REGION Network 20: Total Time Machine
   // ENO of a box is taken as its EN; it also drops when the box reports an error
   "Data_TimeData"."Total Time Machine" := "Data_TimeData"."Mesin Run" + "Data_TimeData"."Mesin Run Baypass" + "Data_TimeData"."Mesin Stop" + "Data_TimeData"."Mesin Error";
   "Data_TODData"."Total Time Machine" := T_CONV(IN := "Data_TimeData"."Total Time Machine");
   "Data_DTLData"."Total Time Machine"[0] := T_COMBINE(IN1 := D#1990-01-01,
                           IN2 := "Data_TODData"."Total Time Machine");
END_REGION

REGION Network 21: % Persen Counter Mesin Terhadap Lama Current Shift
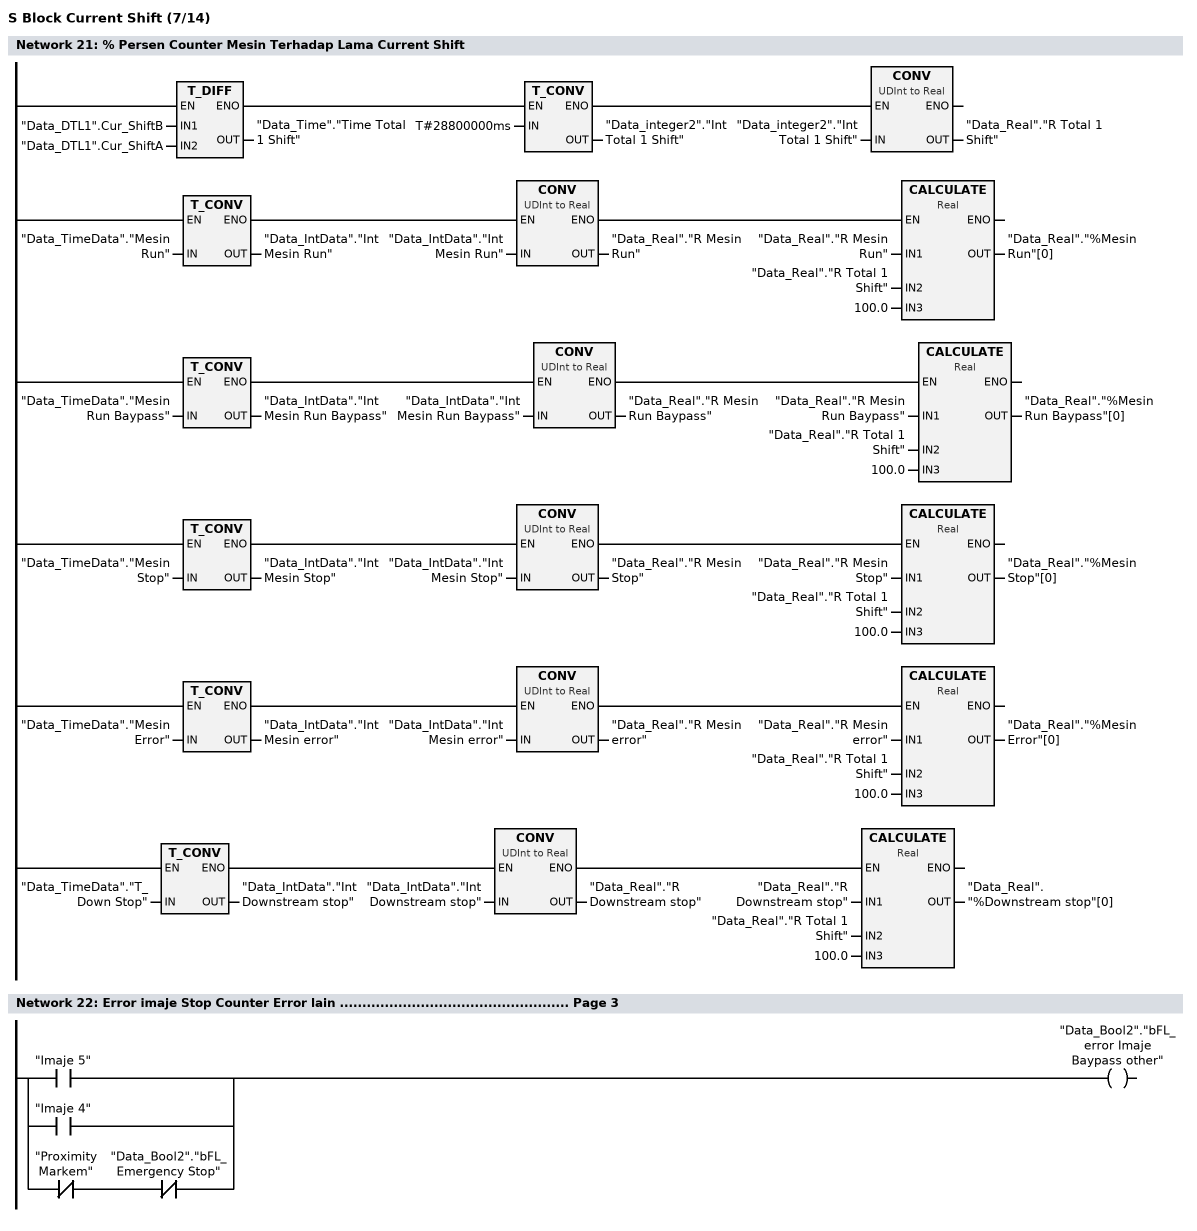
   // ENO of a box is taken as its EN; it also drops when the box reports an error
   "Data_Time"."Time Total 1 Shift" := T_DIFF(IN1 := "Data_DTL1".Cur_ShiftB, IN2 := "Data_DTL1".Cur_ShiftA);
   "Data_integer2"."Int Total 1 Shift" := T_CONV(IN := T#28800000ms);
   "Data_Real"."R Total 1 Shift" := UDINT_TO_REAL("Data_integer2"."Int Total 1 Shift");
   "Data_IntData"."Int Mesin Run" := T_CONV(IN := "Data_TimeData"."Mesin Run");
   "Data_Real"."R Mesin Run" := UDINT_TO_REAL("Data_IntData"."Int Mesin Run");
   "Data_Real"."%Mesin Run"[0] := ("Data_Real"."R Mesin Run"/"Data_Real"."R Total 1 Shift")*100.0;
   "Data_IntData"."Int Mesin Run Baypass" := T_CONV(IN := "Data_TimeData"."Mesin Run Baypass");
   "Data_Real"."R Mesin Run Baypass" := UDINT_TO_REAL("Data_IntData"."Int Mesin Run Baypass");
   "Data_Real"."%Mesin Run Baypass"[0] := ("Data_Real"."R Mesin Run Baypass"/"Data_Real"."R Total 1 Shift")*100.0;
   "Data_IntData"."Int Mesin Stop" := T_CONV(IN := "Data_TimeData"."Mesin Stop");
   "Data_Real"."R Mesin Stop" := UDINT_TO_REAL("Data_IntData"."Int Mesin Stop");
   "Data_Real"."%Mesin Stop"[0] := ("Data_Real"."R Mesin Stop"/"Data_Real"."R Total 1 Shift")*100.0;
   "Data_IntData"."Int Mesin error" := T_CONV(IN := "Data_TimeData"."Mesin Error");
   "Data_Real"."R Mesin error" := UDINT_TO_REAL("Data_IntData"."Int Mesin error");
   "Data_Real"."%Mesin Error"[0] := ("Data_Real"."R Mesin error"/"Data_Real"."R Total 1 Shift")*100.0;
   "Data_IntData"."Int Downstream stop" := T_CONV(IN := "Data_TimeData"."T_Down Stop");
   "Data_Real"."R Downstream stop" := UDINT_TO_REAL("Data_IntData"."Int Downstream stop");
   "Data_Real"."%Downstream stop"[0] := ("Data_Real"."R Downstream stop"/"Data_Real"."R Total 1 Shift")*100.0;
END_REGION

REGION Network 22: Error imaje Stop Counter Error lain ................................................... Page 3
   RUNG wire#powerrail
      Contact( "Imaje 5" )
      wire#w1
      Coil( "Data_Bool2"."bFL_error Imaje Baypass other" )
   END_RUNG
   RUNG wire#powerrail
      Contact( "Imaje 4" )
   END_RUNG wire#w1
   RUNG wire#powerrail
      I_Contact( "Proximity Markem" )
      I_Contact( "Data_Bool2"."bFL_Emergency Stop" )
   END_RUNG wire#w1
   // the same network as SCL:
   "Data_Bool2"."bFL_error Imaje Baypass other" := "Imaje 5" OR "Imaje 4" OR (NOT "Proximity Markem" AND NOT "Data_Bool2"."bFL_Emergency Stop");
END_REGION

REGION Network 23: 1. Counter Imaje System Error
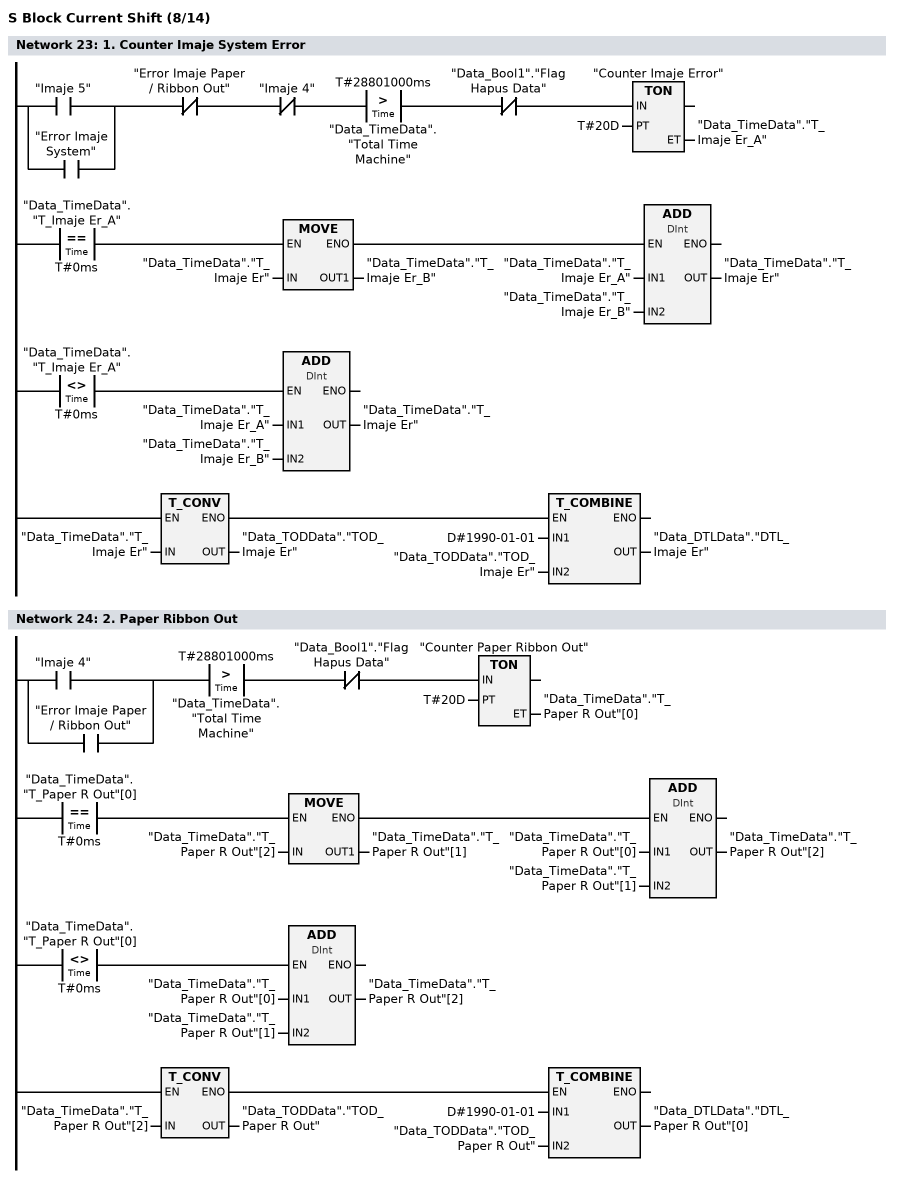
   // ENO of a box is taken as its EN; it also drops when the box reports an error
   "Counter Imaje Error".TON(IN := ("Imaje 5" OR "Error Imaje System") AND NOT "Error Imaje Paper / Ribbon Out" AND NOT "Imaje 4" AND (T#28801000ms > "Data_TimeData"."Total Time Machine") AND NOT "Data_Bool1"."Flag Hapus Data",
                           PT := T#20D,
                           ET => "Data_TimeData"."T_Imaje Er_A");
   IF "Data_TimeData"."T_Imaje Er_A" = T#0ms THEN
       "Data_TimeData"."T_Imaje Er_B" := "Data_TimeData"."T_Imaje Er";
       "Data_TimeData"."T_Imaje Er" := "Data_TimeData"."T_Imaje Er_A" + "Data_TimeData"."T_Imaje Er_B";
   END_IF;
   IF "Data_TimeData"."T_Imaje Er_A" <> T#0ms THEN
       "Data_TimeData"."T_Imaje Er" := "Data_TimeData"."T_Imaje Er_A" + "Data_TimeData"."T_Imaje Er_B";
   END_IF;
   "Data_TODData"."TOD_Imaje Er" := T_CONV(IN := "Data_TimeData"."T_Imaje Er");
   "Data_DTLData"."DTL_Imaje Er" := T_COMBINE(IN1 := D#1990-01-01, IN2 := "Data_TODData"."TOD_Imaje Er");
END_REGION

REGION Network 24: 2. Paper Ribbon Out
   // ENO of a box is taken as its EN; it also drops when the box reports an error
   "Counter Paper Ribbon Out".TON(IN := ("Imaje 4" OR "Error Imaje Paper / Ribbon Out") AND (T#28801000ms > "Data_TimeData"."Total Time Machine") AND NOT "Data_Bool1"."Flag Hapus Data",
                           PT := T#20D,
                           ET => "Data_TimeData"."T_Paper R Out"[0]);
   #_w1 := "Data_TimeData"."T_Paper R Out"[0] = T#0ms;
   IF #_w1 THEN
       "Data_TimeData"."T_Paper R Out"[1] := "Data_TimeData"."T_Paper R Out"[2];
       "Data_TimeData"."T_Paper R Out"[2] := "Data_TimeData"."T_Paper R Out"[0] + "Data_TimeData"."T_Paper R Out"[1];
   END_IF;
   IF "Data_TimeData"."T_Paper R Out"[0] <> T#0ms THEN
       "Data_TimeData"."T_Paper R Out"[2] := "Data_TimeData"."T_Paper R Out"[0] + "Data_TimeData"."T_Paper R Out"[1];
   END_IF;
   "Data_TODData"."TOD_Paper R Out" := T_CONV(IN := "Data_TimeData"."T_Paper R Out"[2]);
   "Data_DTLData"."DTL_Paper R Out"[0] := T_COMBINE(IN1 := D#1990-01-01,
                           IN2 := "Data_TODData"."TOD_Paper R Out");
END_REGION

REGION Network 25: 3. Imaje Not In Position
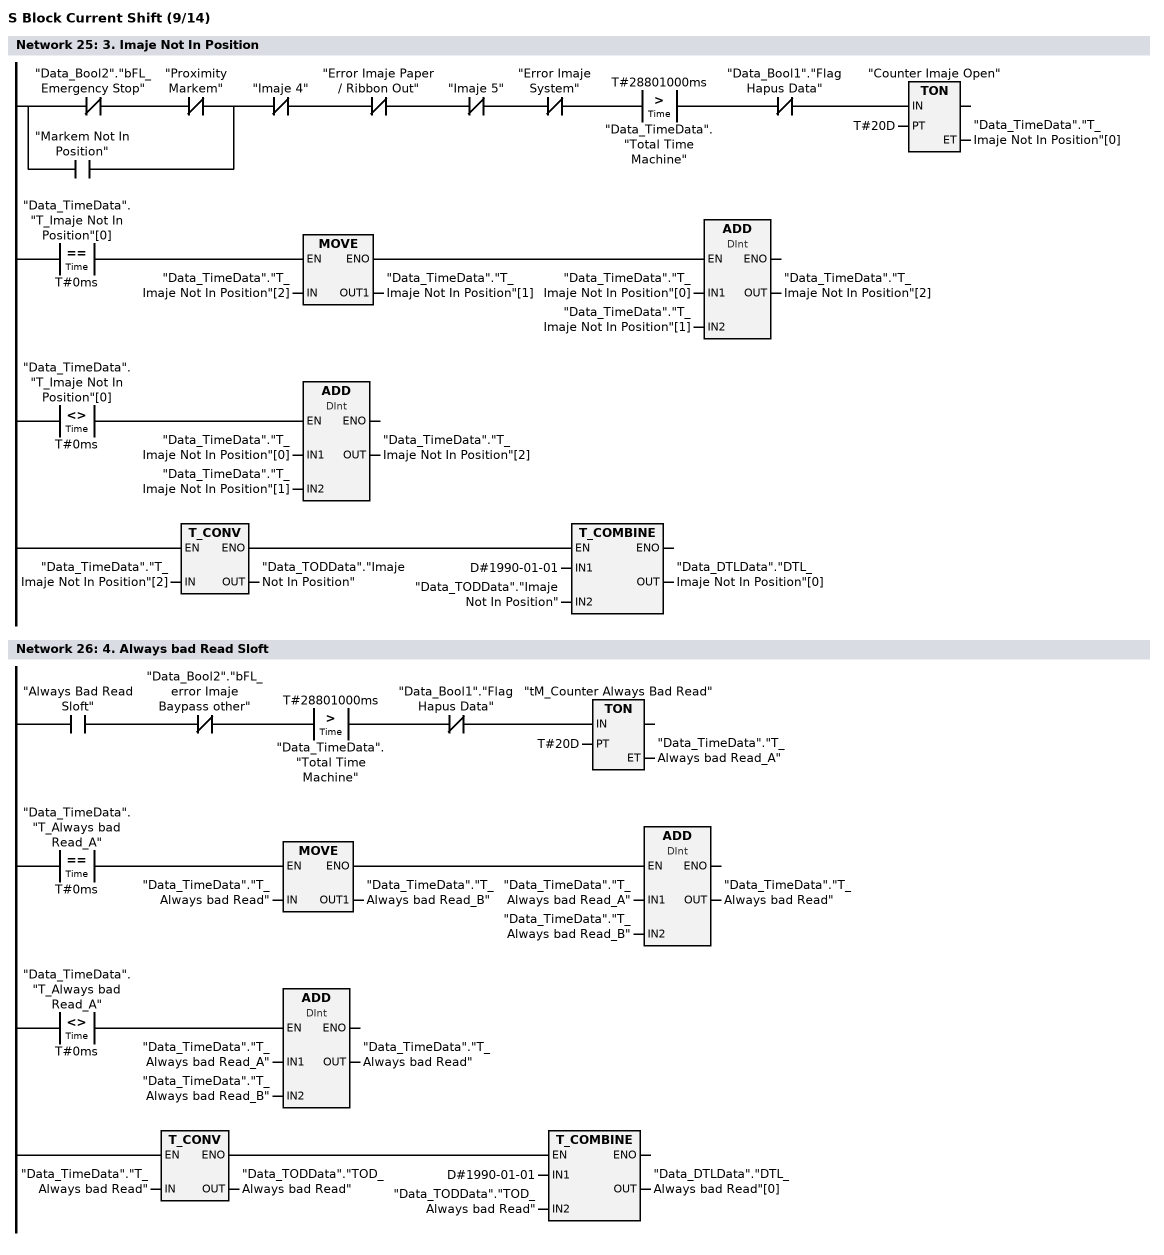
   // ENO of a box is taken as its EN; it also drops when the box reports an error
   "Counter Imaje Open".TON(IN := ((NOT "Data_Bool2"."bFL_Emergency Stop" AND NOT "Proximity Markem") OR "Markem Not In Position") AND NOT "Imaje 4" AND NOT "Error Imaje Paper / Ribbon Out" AND NOT "Imaje 5" AND NOT "Error Imaje System" AND (T#28801000ms > "Data_TimeData"."Total Time Machine") AND NOT "Data_Bool1"."Flag Hapus Data",
                           PT := T#20D,
                           ET => "Data_TimeData"."T_Imaje Not In Position"[0]);
   #_w1 := "Data_TimeData"."T_Imaje Not In Position"[0] = T#0ms;
   IF #_w1 THEN
       "Data_TimeData"."T_Imaje Not In Position"[1] := "Data_TimeData"."T_Imaje Not In Position"[2];
       "Data_TimeData"."T_Imaje Not In Position"[2] := "Data_TimeData"."T_Imaje Not In Position"[0] + "Data_TimeData"."T_Imaje Not In Position"[1];
   END_IF;
   IF "Data_TimeData"."T_Imaje Not In Position"[0] <> T#0ms THEN
       "Data_TimeData"."T_Imaje Not In Position"[2] := "Data_TimeData"."T_Imaje Not In Position"[0] + "Data_TimeData"."T_Imaje Not In Position"[1];
   END_IF;
   "Data_TODData"."Imaje Not In Position" := T_CONV(IN := "Data_TimeData"."T_Imaje Not In Position"[2]);
   "Data_DTLData"."DTL_Imaje Not In Position"[0] := T_COMBINE(IN1 := D#1990-01-01,
                           IN2 := "Data_TODData"."Imaje Not In Position");
END_REGION

REGION Network 26: 4. Always bad Read Sloft
   // ENO of a box is taken as its EN; it also drops when the box reports an error
   "tM_Counter Always Bad Read".TON(IN := "Always Bad Read Sloft" AND NOT "Data_Bool2"."bFL_error Imaje Baypass other" AND (T#28801000ms > "Data_TimeData"."Total Time Machine") AND NOT "Data_Bool1"."Flag Hapus Data",
                           PT := T#20D,
                           ET => "Data_TimeData"."T_Always bad Read_A");
   IF "Data_TimeData"."T_Always bad Read_A" = T#0ms THEN
       "Data_TimeData"."T_Always bad Read_B" := "Data_TimeData"."T_Always bad Read";
       "Data_TimeData"."T_Always bad Read" := "Data_TimeData"."T_Always bad Read_A" + "Data_TimeData"."T_Always bad Read_B";
   END_IF;
   IF "Data_TimeData"."T_Always bad Read_A" <> T#0ms THEN
       "Data_TimeData"."T_Always bad Read" := "Data_TimeData"."T_Always bad Read_A" + "Data_TimeData"."T_Always bad Read_B";
   END_IF;
   "Data_TODData"."TOD_Always bad Read" := T_CONV(IN := "Data_TimeData"."T_Always bad Read");
   "Data_DTLData"."DTL_Always bad Read"[0] := T_COMBINE(IN1 := D#1990-01-01,
                           IN2 := "Data_TODData"."TOD_Always bad Read");
END_REGION

REGION Network 27: 5. Counter Sloft Jammed
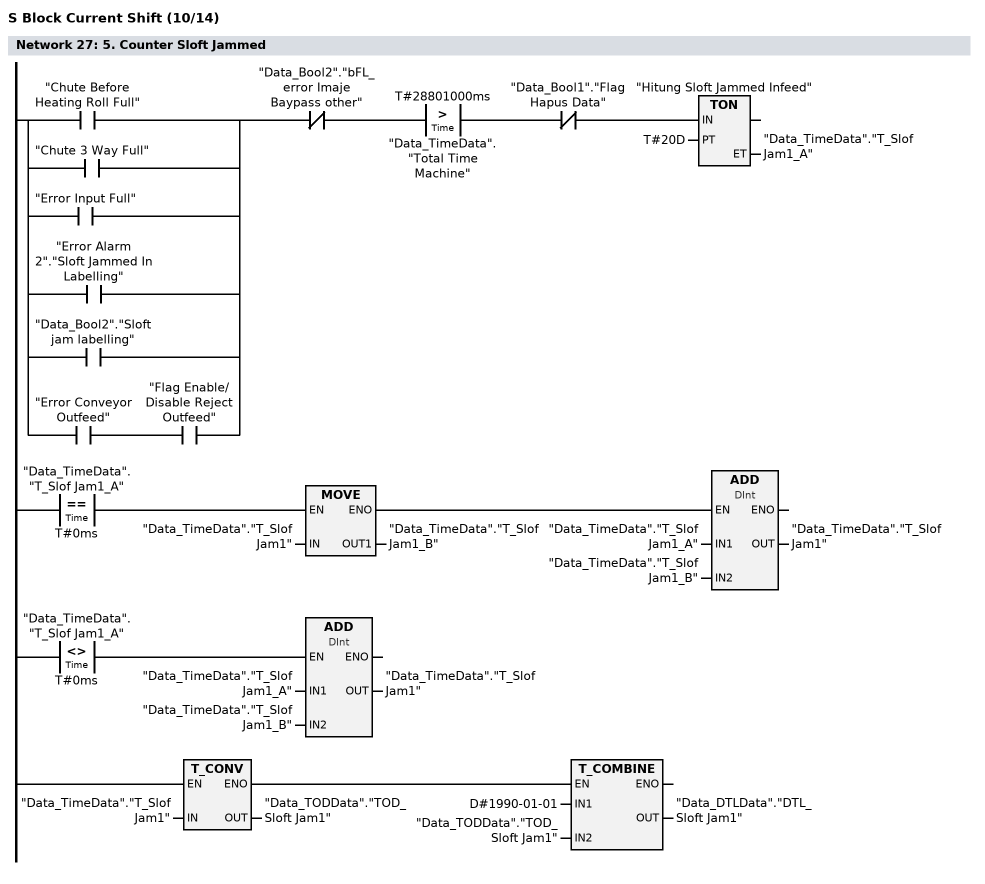
   // ENO of a box is taken as its EN; it also drops when the box reports an error
   "Hitung Sloft Jammed Infeed".TON(IN := ("Chute Before Heating Roll Full" OR "Chute 3 Way Full" OR "Error Input Full" OR "Error Alarm 2"."Sloft Jammed In Labelling" OR "Data_Bool2"."Sloft jam labelling" OR ("Error Conveyor Outfeed" AND "Flag Enable/Disable Reject Outfeed")) AND NOT "Data_Bool2"."bFL_error Imaje Baypass other" AND (T#28801000ms > "Data_TimeData"."Total Time Machine") AND NOT "Data_Bool1"."Flag Hapus Data",
                           PT := T#20D,
                           ET => "Data_TimeData"."T_Slof Jam1_A");
   IF "Data_TimeData"."T_Slof Jam1_A" = T#0ms THEN
       "Data_TimeData"."T_Slof Jam1_B" := "Data_TimeData"."T_Slof Jam1";
       "Data_TimeData"."T_Slof Jam1" := "Data_TimeData"."T_Slof Jam1_A" + "Data_TimeData"."T_Slof Jam1_B";
   END_IF;
   IF "Data_TimeData"."T_Slof Jam1_A" <> T#0ms THEN
       "Data_TimeData"."T_Slof Jam1" := "Data_TimeData"."T_Slof Jam1_A" + "Data_TimeData"."T_Slof Jam1_B";
   END_IF;
   "Data_TODData"."TOD_Sloft Jam1" := T_CONV(IN := "Data_TimeData"."T_Slof Jam1");
   "Data_DTLData"."DTL_Sloft Jam1" := T_COMBINE(IN1 := D#1990-01-01, IN2 := "Data_TODData"."TOD_Sloft Jam1");
END_REGION

REGION Network 28: 6. Counter Pressure Low
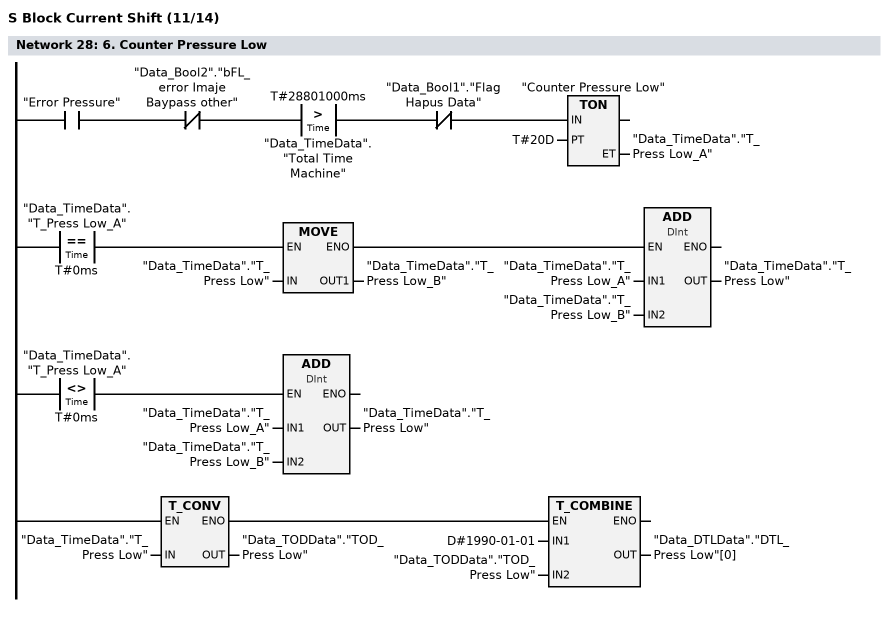
   // ENO of a box is taken as its EN; it also drops when the box reports an error
   "Counter Pressure Low".TON(IN := "Error Pressure" AND NOT "Data_Bool2"."bFL_error Imaje Baypass other" AND (T#28801000ms > "Data_TimeData"."Total Time Machine") AND NOT "Data_Bool1"."Flag Hapus Data",
                           PT := T#20D,
                           ET => "Data_TimeData"."T_Press Low_A");
   IF "Data_TimeData"."T_Press Low_A" = T#0ms THEN
       "Data_TimeData"."T_Press Low_B" := "Data_TimeData"."T_Press Low";
       "Data_TimeData"."T_Press Low" := "Data_TimeData"."T_Press Low_A" + "Data_TimeData"."T_Press Low_B";
   END_IF;
   IF "Data_TimeData"."T_Press Low_A" <> T#0ms THEN
       "Data_TimeData"."T_Press Low" := "Data_TimeData"."T_Press Low_A" + "Data_TimeData"."T_Press Low_B";
   END_IF;
   "Data_TODData"."TOD_Press Low" := T_CONV(IN := "Data_TimeData"."T_Press Low");
   "Data_DTLData"."DTL_Press Low"[0] := T_COMBINE(IN1 := D#1990-01-01, IN2 := "Data_TODData"."TOD_Press Low");
END_REGION

REGION Network 29: 7. Counter RS Pneumatic Error
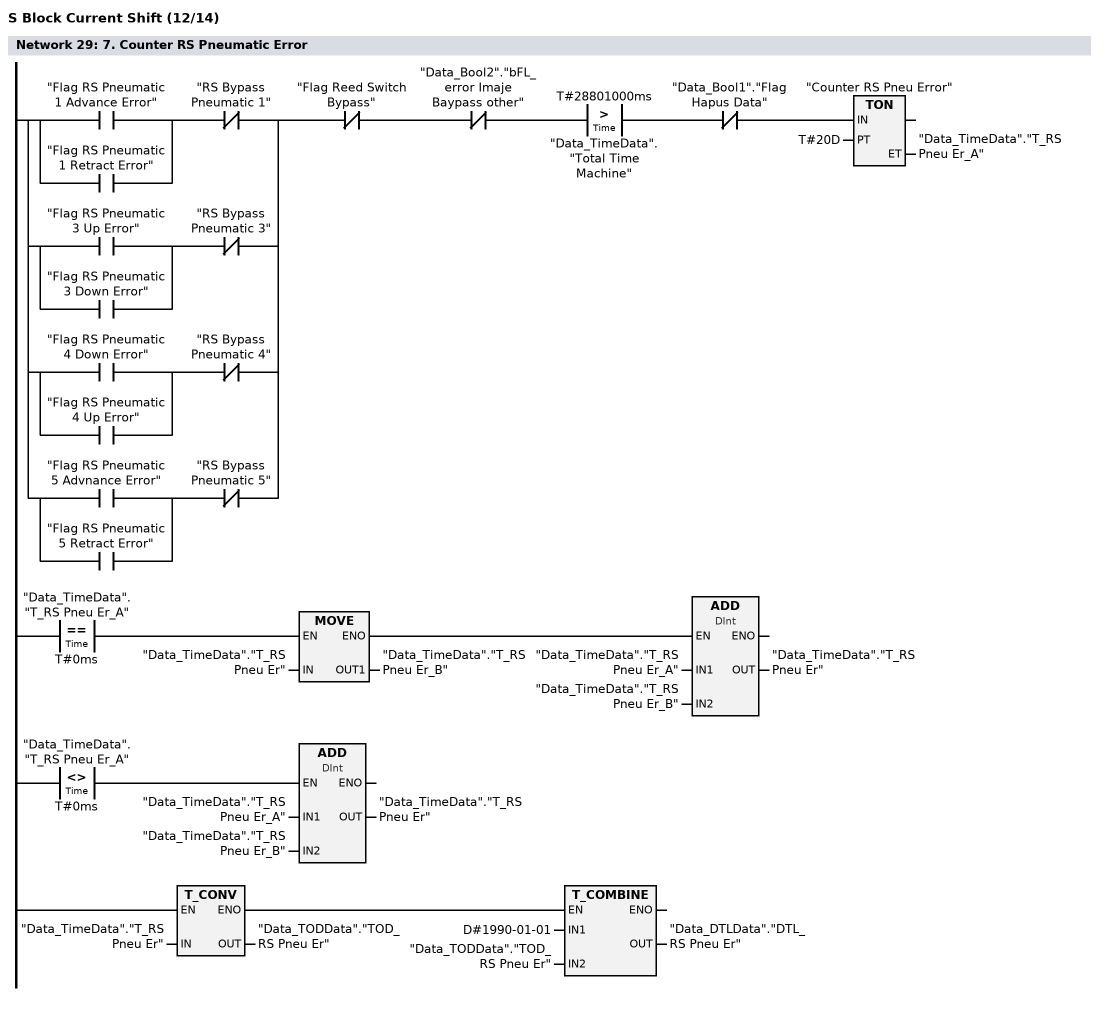
   // ENO of a box is taken as its EN; it also drops when the box reports an error
   "Counter RS Pneu Error".TON(IN := ((("Flag RS Pneumatic 1 Advance Error" OR "Flag RS Pneumatic 1 Retract Error") AND NOT "RS Bypass Pneumatic 1") OR (("Flag RS Pneumatic 3 Up Error" OR "Flag RS Pneumatic 3 Down Error") AND NOT "RS Bypass Pneumatic 3") OR (("Flag RS Pneumatic 4 Down Error" OR "Flag RS Pneumatic 4 Up Error") AND NOT "RS Bypass Pneumatic 4") OR (("Flag RS Pneumatic 5 Advnance Error" OR "Flag RS Pneumatic 5 Retract Error") AND NOT "RS Bypass Pneumatic 5")) AND NOT "Flag Reed Switch Bypass" AND NOT "Data_Bool2"."bFL_error Imaje Baypass other" AND (T#28801000ms > "Data_TimeData"."Total Time Machine") AND NOT "Data_Bool1"."Flag Hapus Data",
                           PT := T#20D,
                           ET => "Data_TimeData"."T_RS Pneu Er_A");
   IF "Data_TimeData"."T_RS Pneu Er_A" = T#0ms THEN
       "Data_TimeData"."T_RS Pneu Er_B" := "Data_TimeData"."T_RS Pneu Er";
       "Data_TimeData"."T_RS Pneu Er" := "Data_TimeData"."T_RS Pneu Er_A" + "Data_TimeData"."T_RS Pneu Er_B";
   END_IF;
   IF "Data_TimeData"."T_RS Pneu Er_A" <> T#0ms THEN
       "Data_TimeData"."T_RS Pneu Er" := "Data_TimeData"."T_RS Pneu Er_A" + "Data_TimeData"."T_RS Pneu Er_B";
   END_IF;
   "Data_TODData"."TOD_RS Pneu Er" := T_CONV(IN := "Data_TimeData"."T_RS Pneu Er");
   "Data_DTLData"."DTL_RS Pneu Er" := T_COMBINE(IN1 := D#1990-01-01, IN2 := "Data_TODData"."TOD_RS Pneu Er");
END_REGION

REGION Network 30: 8. Counter Door open error
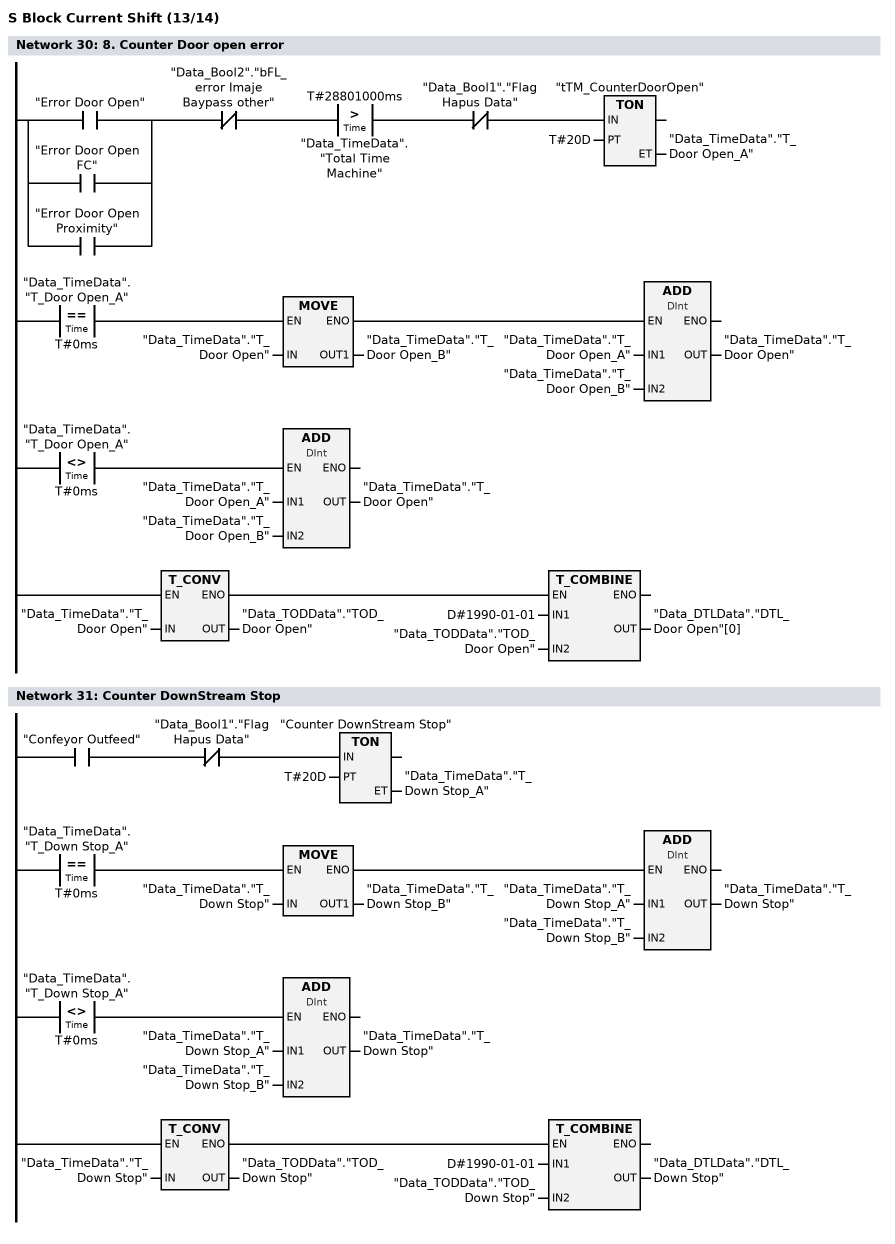
   // ENO of a box is taken as its EN; it also drops when the box reports an error
   "tTM_CounterDoorOpen".TON(IN := ("Error Door Open" OR "Error Door Open FC" OR "Error Door Open Proximity") AND NOT "Data_Bool2"."bFL_error Imaje Baypass other" AND (T#28801000ms > "Data_TimeData"."Total Time Machine") AND NOT "Data_Bool1"."Flag Hapus Data",
                           PT := T#20D,
                           ET => "Data_TimeData"."T_Door Open_A");
   IF "Data_TimeData"."T_Door Open_A" = T#0ms THEN
       "Data_TimeData"."T_Door Open_B" := "Data_TimeData"."T_Door Open";
       "Data_TimeData"."T_Door Open" := "Data_TimeData"."T_Door Open_A" + "Data_TimeData"."T_Door Open_B";
   END_IF;
   IF "Data_TimeData"."T_Door Open_A" <> T#0ms THEN
       "Data_TimeData"."T_Door Open" := "Data_TimeData"."T_Door Open_A" + "Data_TimeData"."T_Door Open_B";
   END_IF;
   "Data_TODData"."TOD_Door Open" := T_CONV(IN := "Data_TimeData"."T_Door Open");
   "Data_DTLData"."DTL_Door Open"[0] := T_COMBINE(IN1 := D#1990-01-01, IN2 := "Data_TODData"."TOD_Door Open");
END_REGION

REGION Network 31: Counter DownStream Stop
   // ENO of a box is taken as its EN; it also drops when the box reports an error
   "Counter DownStream Stop".TON(IN := "Confeyor Outfeed" AND NOT "Data_Bool1"."Flag Hapus Data",
                           PT := T#20D,
                           ET => "Data_TimeData"."T_Down Stop_A");
   IF "Data_TimeData"."T_Down Stop_A" = T#0ms THEN
       "Data_TimeData"."T_Down Stop_B" := "Data_TimeData"."T_Down Stop";
       "Data_TimeData"."T_Down Stop" := "Data_TimeData"."T_Down Stop_A" + "Data_TimeData"."T_Down Stop_B";
   END_IF;
   IF "Data_TimeData"."T_Down Stop_A" <> T#0ms THEN
       "Data_TimeData"."T_Down Stop" := "Data_TimeData"."T_Down Stop_A" + "Data_TimeData"."T_Down Stop_B";
   END_IF;
   "Data_TODData"."TOD_Down Stop" := T_CONV(IN := "Data_TimeData"."T_Down Stop");
   "Data_DTLData"."DTL_Down Stop" := T_COMBINE(IN1 := D#1990-01-01, IN2 := "Data_TODData"."TOD_Down Stop");
END_REGION

REGION Network 32: Total Error
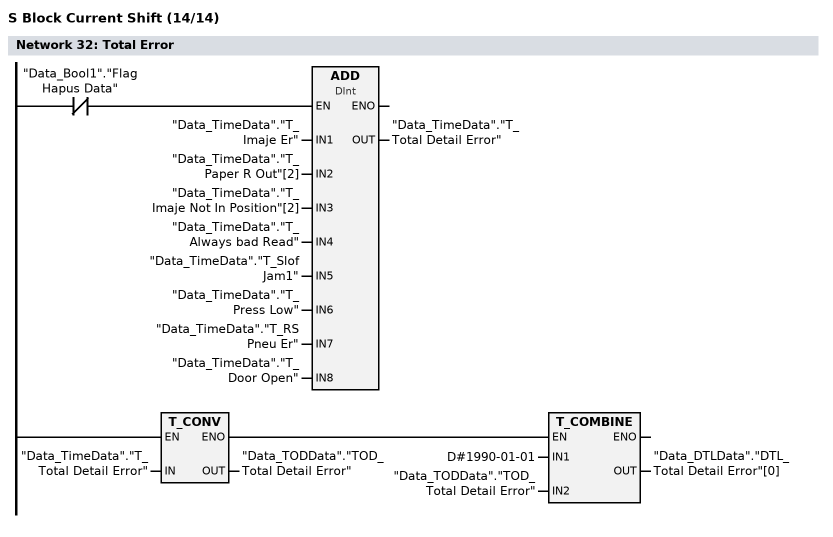
   // ENO of a box is taken as its EN; it also drops when the box reports an error
   IF NOT "Data_Bool1"."Flag Hapus Data" THEN
       "Data_TimeData"."T_Total Detail Error" := "Data_TimeData"."T_Imaje Er" + "Data_TimeData"."T_Paper R Out"[2] + "Data_TimeData"."T_Imaje Not In Position"[2] + "Data_TimeData"."T_Always bad Read" + "Data_TimeData"."T_Slof Jam1" + "Data_TimeData"."T_Press Low" + "Data_TimeData"."T_RS Pneu Er" + "Data_TimeData"."T_Door Open";
   END_IF;
   "Data_TODData"."TOD_Total Detail Error" := T_CONV(IN := "Data_TimeData"."T_Total Detail Error");
   "Data_DTLData"."DTL_Total Detail Error"[0] := T_COMBINE(IN1 := D#1990-01-01,
                           IN2 := "Data_TODData"."TOD_Total Detail Error");
END_REGION
END_FUNCTION_BLOCK

FUNCTION_BLOCK "Block Labeling"   // FB5, LAD
{ S7_Optimized_Access := 'TRUE' }
VERSION : 0.1
   VAR_TEMP   // added for the SCL form of the ladder/FBD networks
      _w1 : Bool;
      _w2 : Bool;
      _w3 : Bool;
      _w4 : Bool;
   END_VAR
BEGIN

REGION Network 1: By pass ON
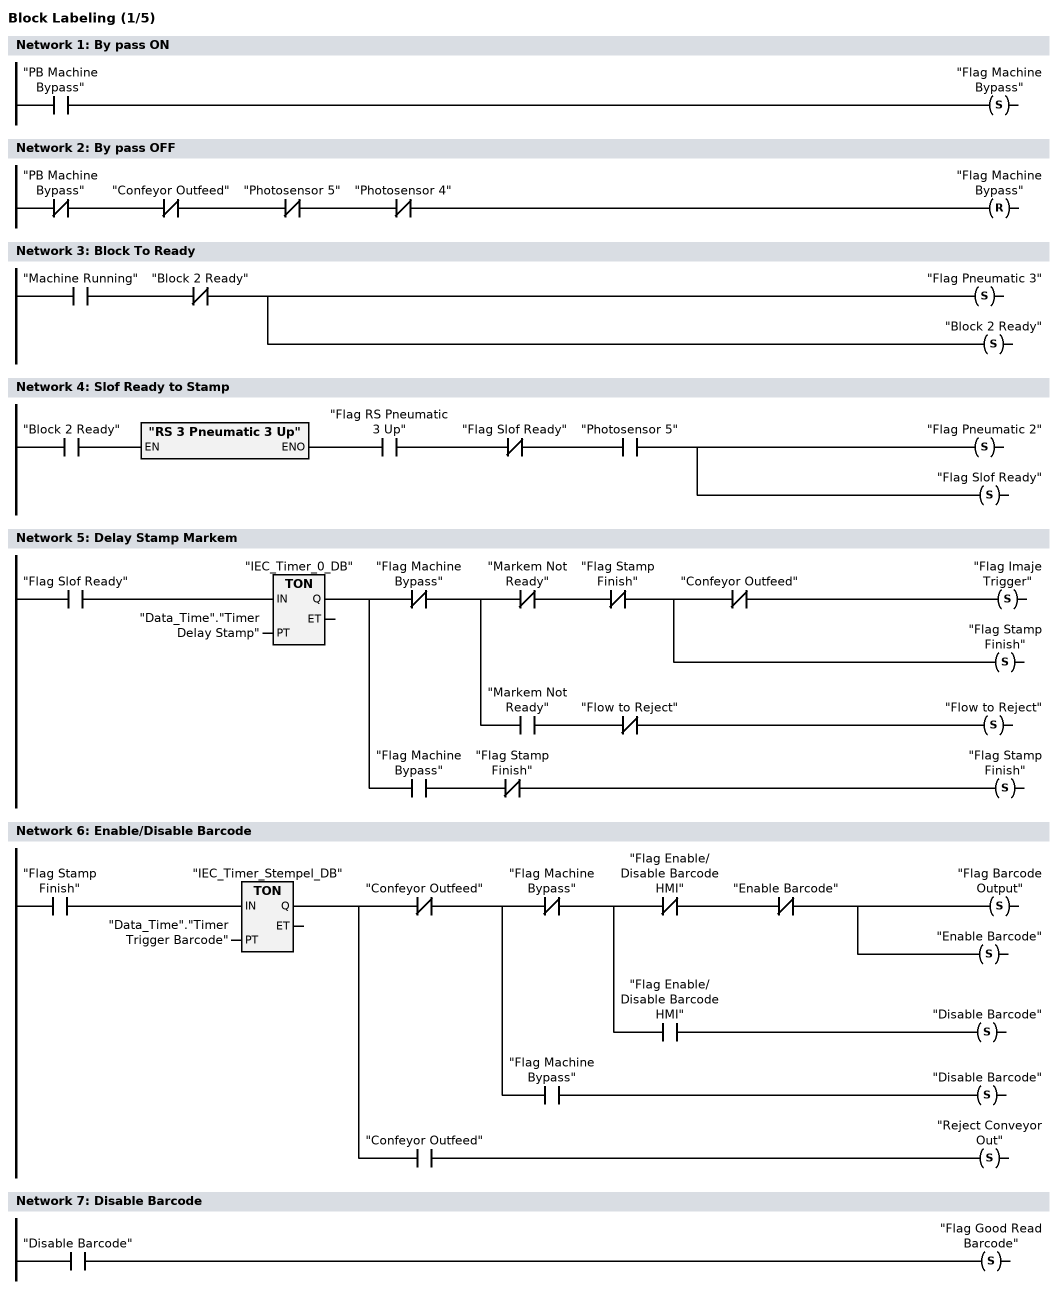
   RUNG wire#powerrail
      Contact( "PB Machine Bypass" )
      S_Coil( "Flag Machine Bypass" )
   END_RUNG
   // the same network as SCL:
   IF "PB Machine Bypass" THEN "Flag Machine Bypass" := TRUE; END_IF;
END_REGION

REGION Network 2: By pass OFF
   RUNG wire#powerrail
      I_Contact( "PB Machine Bypass" )
      I_Contact( "Confeyor Outfeed" )
      I_Contact( "Photosensor 5" )
      I_Contact( "Photosensor 4" )
      R_Coil( "Flag Machine Bypass" )
   END_RUNG
   // the same network as SCL:
   IF NOT "PB Machine Bypass" AND NOT "Confeyor Outfeed" AND NOT "Photosensor 5" AND NOT "Photosensor 4" THEN
       "Flag Machine Bypass" := FALSE;
   END_IF;
END_REGION

REGION Network 3: Block To Ready
   RUNG wire#powerrail
      Contact( "Machine Running" )
      I_Contact( "Block 2 Ready" )
      wire#w1
      S_Coil( "Flag Pneumatic 3" )
   END_RUNG
   RUNG wire#w1
      S_Coil( "Block 2 Ready" )
   END_RUNG
   // the same network as SCL:
   IF "Machine Running" AND NOT "Block 2 Ready" THEN
       "Flag Pneumatic 3" := TRUE;
       "Block 2 Ready" := TRUE;
   END_IF;
END_REGION

REGION Network 4: Slof Ready to Stamp
   RUNG wire#powerrail
      Contact( "Block 2 Ready" )
      "RS 3 Pneumatic 3 Up"()
      Contact( "Flag RS Pneumatic 3 Up" )
      I_Contact( "Flag Slof Ready" )
      Contact( "Photosensor 5" )
      wire#w1
      S_Coil( "Flag Pneumatic 2" )
   END_RUNG
   RUNG wire#w1
      S_Coil( "Flag Slof Ready" )
   END_RUNG
   // the same network as SCL:
   "RS 3 Pneumatic 3 Up"(EN := "Block 2 Ready", ENO => #_w1);
   IF #_w1 AND "Flag RS Pneumatic 3 Up" AND NOT "Flag Slof Ready" AND "Photosensor 5" THEN
       "Flag Pneumatic 2" := TRUE;
       "Flag Slof Ready" := TRUE;
   END_IF;
END_REGION

REGION Network 5: Delay Stamp Markem
   "IEC_Timer_0_DB".TON(IN := "Flag Slof Ready", PT := "Data_Time"."Timer Delay Stamp");
   #_w1 := "IEC_Timer_0_DB".Q AND NOT "Flag Machine Bypass";
   #_w2 := #_w1 AND NOT "Markem Not Ready" AND NOT "Flag Stamp Finish";
   IF #_w2 AND NOT "Confeyor Outfeed" THEN "Flag Imaje Trigger" := TRUE; END_IF;
   IF #_w2 THEN "Flag Stamp Finish" := TRUE; END_IF;
   IF #_w1 AND "Markem Not Ready" AND NOT "Flow to Reject" THEN "Flow to Reject" := TRUE; END_IF;
   IF "IEC_Timer_0_DB".Q AND "Flag Machine Bypass" AND NOT "Flag Stamp Finish" THEN
       "Flag Stamp Finish" := TRUE;
   END_IF;
END_REGION

REGION Network 6: Enable/Disable Barcode
   "IEC_Timer_Stempel_DB".TON(IN := "Flag Stamp Finish", PT := "Data_Time"."Timer Trigger Barcode");
   #_w1 := "IEC_Timer_Stempel_DB".Q AND NOT "Confeyor Outfeed";
   #_w2 := #_w1 AND NOT "Flag Machine Bypass";
   IF #_w2 AND NOT "Flag Enable/Disable Barcode HMI" AND NOT "Enable Barcode" THEN
       "Flag Barcode Output" := TRUE;
       "Enable Barcode" := TRUE;
   END_IF;
   IF #_w2 AND "Flag Enable/Disable Barcode HMI" THEN "Disable Barcode" := TRUE; END_IF;
   IF #_w1 AND "Flag Machine Bypass" THEN "Disable Barcode" := TRUE; END_IF;
   IF "IEC_Timer_Stempel_DB".Q AND "Confeyor Outfeed" THEN "Reject Conveyor Out" := TRUE; END_IF;
END_REGION

REGION Network 7: Disable Barcode
   RUNG wire#powerrail
      Contact( "Disable Barcode" )
      S_Coil( "Flag Good Read Barcode" )
   END_RUNG
   // the same network as SCL:
   IF "Disable Barcode" THEN "Flag Good Read Barcode" := TRUE; END_IF;
END_REGION

REGION Network 8: Check Barcode